REGION Network 77: Status signals
   RUNG wire#powerrail
      Contact( #TMP_xAlwaysON )
      wire#w1
      Contact( #STC_tPZD_OpCLLoop.tR.tZSW1.x0 )
      Coil( #STC_tUSER_DATA.tR.xReadyfForSwitchOn )
   END_RUNG
   RUNG wire#w1
      Contact( #STC_tPZD_OpCLLoop.tR.tZSW1.x1 )
      Contact( #STC_tPZD_OpCLLoop.tR.tZSW1.x2 )
      Coil( #STC_tUSER_DATA.tR.xReadyToMove )
   END_RUNG
   RUNG wire#w1
      Contact( #STC_tPZD_OpCLLoop.tR.tZSW1.x1 )
      Contact( #STC_tPZD_OpCLLoop.tR.tZSW1.x10 )
      Coil( #OUT_xFeedback )
   END_RUNG
   RUNG wire#w1
      Contact( #STC_tPZD_OpCLLoop.tR.tZSW1.x3 )
      wire#w2
      Coil( #OUT_xFaultPresent )
   END_RUNG
   RUNG wire#w1
      { S7_Templates := "SrcType := Int" } NE_Contact(in1 := #OUT_iRetVal, in2 := 0)
   END_RUNG wire#w2
   RUNG wire#w1
      Contact( #STC_tPZD_OpCLLoop.tR.tZSW1.x7 )
      Coil( #STC_tUSER_DATA.tR.xAlarmPresent )
   END_RUNG
   // the same network as SCL:
   #STC_tUSER_DATA.tR.xReadyfForSwitchOn := #TMP_xAlwaysON AND #STC_tPZD_OpCLLoop.tR.tZSW1.x0;
   #STC_tUSER_DATA.tR.xReadyToMove := #TMP_xAlwaysON AND #STC_tPZD_OpCLLoop.tR.tZSW1.x1 AND #STC_tPZD_OpCLLoop.tR.tZSW1.x2;
   #OUT_xFeedback := #TMP_xAlwaysON AND #STC_tPZD_OpCLLoop.tR.tZSW1.x1 AND #STC_tPZD_OpCLLoop.tR.tZSW1.x10;
   #OUT_xFaultPresent := #TMP_xAlwaysON AND (#STC_tPZD_OpCLLoop.tR.tZSW1.x3 OR (#OUT_iRetVal <> 0));
   #STC_tUSER_DATA.tR.xAlarmPresent := #TMP_xAlwaysON AND #STC_tPZD_OpCLLoop.tR.tZSW1.x7;
END_REGION

REGION Network 78: Status values
   RUNG wire#powerrail
      Contact( #TMP_xAlwaysON )
      wire#w1
      { S7_Templates := "[SrcType := DInt, DestType := Real]"; S7_GenerateENO := "TRUE" } Convert(in := #STC_tSYS_DATA.dMaxSpeed_rpm, out => #TMP_r)
      { S7_Templates := "SrcType := Real"; S7_GenerateENO := "TRUE" } Div(in1 := 16384.0, in2 := #TMP_r, out => #TMP_r)
   END_RUNG
   RUNG wire#w1
      { S7_Templates := "[SrcType := Int, DestType := DInt]"; S7_GenerateENO := "TRUE" } Convert(in := #STC_tPZD_OpCLLoop.tR.iNIST_A, out => #TMP_d)
      { S7_Templates := "[SrcType := DInt, DestType := Real]"; S7_GenerateENO := "TRUE" } Convert(in := #TMP_d, out => #TMP_rActualSpeed)
   END_RUNG
   RUNG wire#w1
      { S7_Templates := "SrcType := Real"; S7_GenerateENO := "TRUE" } Div(in1 := #TMP_rActualSpeed, in2 := #TMP_r, out => #TMP_rActualSpeed)
      { S7_Templates := "SrcType := Real"; S7_GenerateENO := "TRUE" } Mul(in1 := #TMP_rActualSpeed, in2 := #STC_tSYS_DATA.rK_rpm_mmMin, out => #TMP_rActualSpeed)
      { S7_Templates := "[SrcType := Real, DestType := DInt]"; S7_GenerateENO := "TRUE" } Trunc(in := #TMP_rActualSpeed, out => #STC_tUSER_DATA.tR.dActualSpeed_mm_min)
   END_RUNG
   // the same network as SCL:
   // ENO of a box is taken as its EN; it also drops when the box reports an error
   IF #TMP_xAlwaysON THEN
       #TMP_r := DINT_TO_REAL(#STC_tSYS_DATA.dMaxSpeed_rpm);
       #TMP_r := 16384.0 / #TMP_r;
       #TMP_d := INT_TO_DINT(#STC_tPZD_OpCLLoop.tR.iNIST_A);
       #TMP_rActualSpeed := DINT_TO_REAL(#TMP_d);
       #TMP_rActualSpeed := #TMP_rActualSpeed / #TMP_r;
       #TMP_rActualSpeed := #TMP_rActualSpeed * #STC_tSYS_DATA.rK_rpm_mmMin;
       #STC_tUSER_DATA.tR.dActualSpeed_mm_min := TRUNC(#TMP_rActualSpeed);
   END_IF;
END_REGION

REGION Network 79: #####_STATUSES_#####
END_REGION

REGION Network 80: #####_ALARMS_#####
END_REGION

REGION Network 81: Reset faults
   RUNG wire#powerrail
      Contact( #STC_tPZD_OpCLLoop.tR.tZSW1.x3 )
      Contact( #IN_xResetFaults )
      Coil( #STC_tPZD_OpCLLoop.tW.tSTW1.x7 )
   END_RUNG
   // the same network as SCL:
   #STC_tPZD_OpCLLoop.tW.tSTW1.x7 := #STC_tPZD_OpCLLoop.tR.tZSW1.x3 AND #IN_xResetFaults;
END_REGION

REGION Network 82: Fault messages
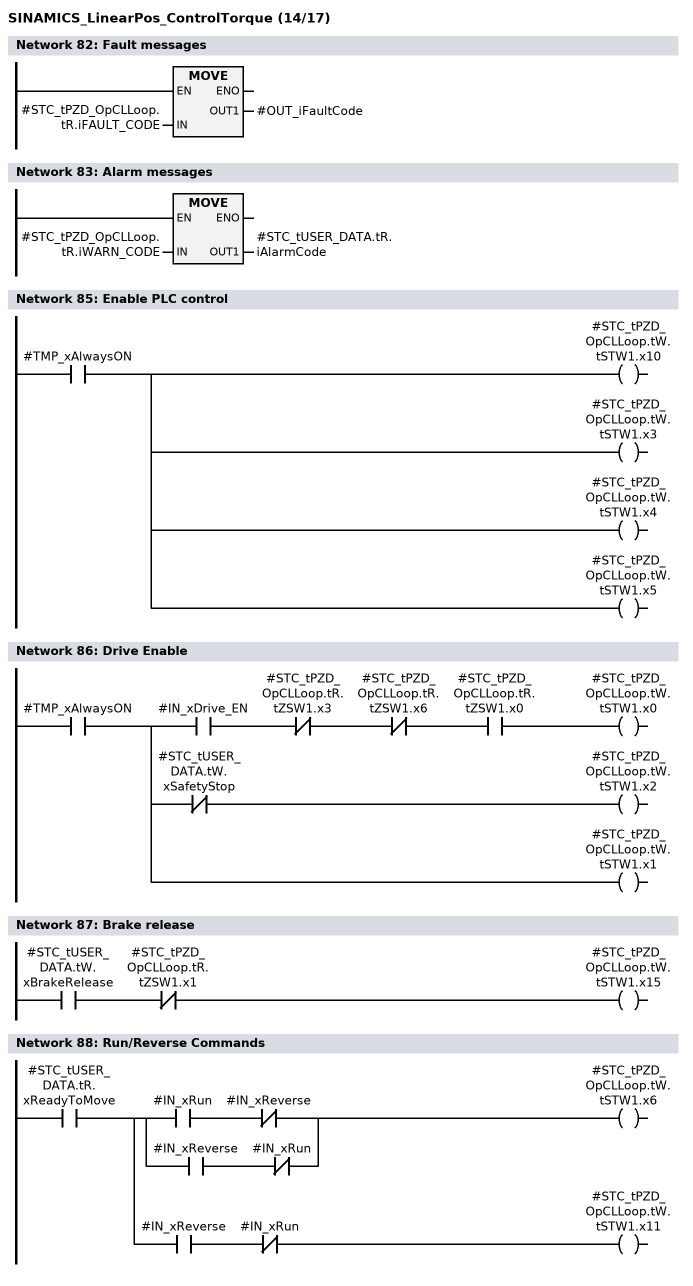
   RUNG wire#powerrail
      { S7_GenerateENO := "TRUE" } Move(in := #STC_tPZD_OpCLLoop.tR.iFAULT_CODE, out1 => #OUT_iFaultCode)
   END_RUNG
   // the same network as SCL:
   #OUT_iFaultCode := #STC_tPZD_OpCLLoop.tR.iFAULT_CODE;
END_REGION

REGION Network 83: Alarm messages
   RUNG wire#powerrail
      { S7_GenerateENO := "TRUE" } Move(in := #STC_tPZD_OpCLLoop.tR.iWARN_CODE, out1 => #STC_tUSER_DATA.tR.iAlarmCode)
   END_RUNG
   // the same network as SCL:
   #STC_tUSER_DATA.tR.iAlarmCode := #STC_tPZD_OpCLLoop.tR.iWARN_CODE;
END_REGION

REGION Network 84: #####_PHASES_&_LOGICS_#####
END_REGION

REGION Network 85: Enable PLC control
   RUNG wire#powerrail
      Contact( #TMP_xAlwaysON )
      wire#w1
      Coil( #STC_tPZD_OpCLLoop.tW.tSTW1.x10 )
   END_RUNG
   RUNG wire#w1
      Coil( #STC_tPZD_OpCLLoop.tW.tSTW1.x3 )
   END_RUNG
   RUNG wire#w1
      Coil( #STC_tPZD_OpCLLoop.tW.tSTW1.x4 )
   END_RUNG
   RUNG wire#w1
      Coil( #STC_tPZD_OpCLLoop.tW.tSTW1.x5 )
   END_RUNG
   // the same network as SCL:
   #STC_tPZD_OpCLLoop.tW.tSTW1.x10 := #TMP_xAlwaysON;
   #STC_tPZD_OpCLLoop.tW.tSTW1.x3 := #TMP_xAlwaysON;
   #STC_tPZD_OpCLLoop.tW.tSTW1.x4 := #TMP_xAlwaysON;
   #STC_tPZD_OpCLLoop.tW.tSTW1.x5 := #TMP_xAlwaysON;
END_REGION

REGION Network 86: Drive Enable
   RUNG wire#powerrail
      Contact( #TMP_xAlwaysON )
      wire#w1
      Contact( #IN_xDrive_EN )
      I_Contact( #STC_tPZD_OpCLLoop.tR.tZSW1.x3 )
      I_Contact( #STC_tPZD_OpCLLoop.tR.tZSW1.x6 )
      Contact( #STC_tPZD_OpCLLoop.tR.tZSW1.x0 )
      Coil( #STC_tPZD_OpCLLoop.tW.tSTW1.x0 )
   END_RUNG
   RUNG wire#w1
      I_Contact( #STC_tUSER_DATA.tW.xSafetyStop )
      Coil( #STC_tPZD_OpCLLoop.tW.tSTW1.x2 )
   END_RUNG
   RUNG wire#w1
      Coil( #STC_tPZD_OpCLLoop.tW.tSTW1.x1 )
   END_RUNG
   // the same network as SCL:
   #STC_tPZD_OpCLLoop.tW.tSTW1.x0 := #TMP_xAlwaysON AND #IN_xDrive_EN AND NOT #STC_tPZD_OpCLLoop.tR.tZSW1.x3 AND NOT #STC_tPZD_OpCLLoop.tR.tZSW1.x6 AND #STC_tPZD_OpCLLoop.tR.tZSW1.x0;
   #STC_tPZD_OpCLLoop.tW.tSTW1.x2 := #TMP_xAlwaysON AND NOT #STC_tUSER_DATA.tW.xSafetyStop;
   #STC_tPZD_OpCLLoop.tW.tSTW1.x1 := #TMP_xAlwaysON;
END_REGION

REGION Network 87: Brake release
   RUNG wire#powerrail
      Contact( #STC_tUSER_DATA.tW.xBrakeRelease )
      I_Contact( #STC_tPZD_OpCLLoop.tR.tZSW1.x1 )
      Coil( #STC_tPZD_OpCLLoop.tW.tSTW1.x15 )
   END_RUNG
   // the same network as SCL:
   #STC_tPZD_OpCLLoop.tW.tSTW1.x15 := #STC_tUSER_DATA.tW.xBrakeRelease AND NOT #STC_tPZD_OpCLLoop.tR.tZSW1.x1;
END_REGION

REGION Network 88: Run/Reverse Commands
   RUNG wire#powerrail
      Contact( #STC_tUSER_DATA.tR.xReadyToMove )
      wire#w1
      Contact( #IN_xRun )
      I_Contact( #IN_xReverse )
      wire#w2
      Coil( #STC_tPZD_OpCLLoop.tW.tSTW1.x6 )
   END_RUNG
   RUNG wire#w1
      Contact( #IN_xReverse )
      I_Contact( #IN_xRun )
   END_RUNG wire#w2
   RUNG wire#w1
      Contact( #IN_xReverse )
      I_Contact( #IN_xRun )
      Coil( #STC_tPZD_OpCLLoop.tW.tSTW1.x11 )
   END_RUNG
   // the same network as SCL:
   #STC_tPZD_OpCLLoop.tW.tSTW1.x6 := #STC_tUSER_DATA.tR.xReadyToMove AND ((#IN_xRun AND NOT #IN_xReverse) OR (#IN_xReverse AND NOT #IN_xRun));
   #STC_tPZD_OpCLLoop.tW.tSTW1.x11 := #STC_tUSER_DATA.tR.xReadyToMove AND #IN_xReverse AND NOT #IN_xRun;
END_REGION

REGION Network 89: #####_PARAMETERS_#####
END_REGION

REGION Network 90: Speed
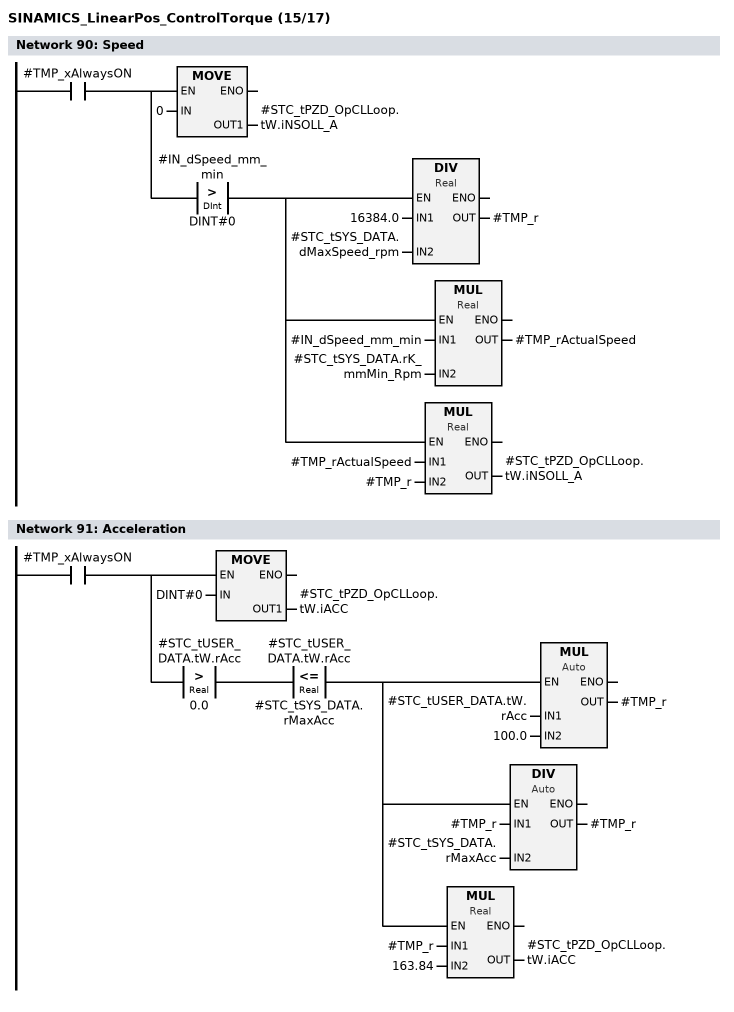
   RUNG wire#powerrail
      Contact( #TMP_xAlwaysON )
      wire#w1
      Move(in := 0, out1 => #STC_tPZD_OpCLLoop.tW.iNSOLL_A)
   END_RUNG
   RUNG wire#w1
      { S7_Templates := "SrcType := DInt" } GT_Contact(in1 := #IN_dSpeed_mm_min, in2 := DINT#0)
      wire#w2
      { S7_Templates := "SrcType := Real" } Div(in1 := 16384.0, in2 := #STC_tSYS_DATA.dMaxSpeed_rpm, out => #TMP_r)
   END_RUNG
   RUNG wire#w2
      { S7_Templates := "SrcType := Real" } Mul(in1 := #IN_dSpeed_mm_min, in2 := #STC_tSYS_DATA.rK_mmMin_Rpm, out => #TMP_rActualSpeed)
   END_RUNG
   RUNG wire#w2
      { S7_Templates := "SrcType := Real" } Mul(in1 := #TMP_rActualSpeed, in2 := #TMP_r, out => #STC_tPZD_OpCLLoop.tW.iNSOLL_A)
   END_RUNG
   // the same network as SCL:
   IF #TMP_xAlwaysON THEN #STC_tPZD_OpCLLoop.tW.iNSOLL_A := 0; END_IF;
   IF #TMP_xAlwaysON AND (#IN_dSpeed_mm_min > DINT#0) THEN
       #TMP_r := 16384.0 / #STC_tSYS_DATA.dMaxSpeed_rpm;
       #TMP_rActualSpeed := #IN_dSpeed_mm_min * #STC_tSYS_DATA.rK_mmMin_Rpm;
       #STC_tPZD_OpCLLoop.tW.iNSOLL_A := #TMP_rActualSpeed * #TMP_r;
   END_IF;
END_REGION

REGION Network 91: Acceleration
   RUNG wire#powerrail
      Contact( #TMP_xAlwaysON )
      wire#w1
      Move(in := DINT#0, out1 => #STC_tPZD_OpCLLoop.tW.iACC)
   END_RUNG
   RUNG wire#w1
      { S7_Templates := "SrcType := Real" } GT_Contact(in1 := #STC_tUSER_DATA.tW.rAcc, in2 := 0.0)
      { S7_Templates := "SrcType := Real" } LE_Contact(in1 := #STC_tUSER_DATA.tW.rAcc, in2 := #STC_tSYS_DATA.rMaxAcc)
      wire#w2
      Mul(in1 := #STC_tUSER_DATA.tW.rAcc, in2 := 100.0, out => #TMP_r)
   END_RUNG
   RUNG wire#w2
      Div(in1 := #TMP_r, in2 := #STC_tSYS_DATA.rMaxAcc, out => #TMP_r)
   END_RUNG
   RUNG wire#w2
      { S7_Templates := "SrcType := Real" } Mul(in1 := #TMP_r, in2 := 163.84, out => #STC_tPZD_OpCLLoop.tW.iACC)
   END_RUNG
   // the same network as SCL:
   IF #TMP_xAlwaysON THEN #STC_tPZD_OpCLLoop.tW.iACC := DINT#0; END_IF;
   IF #TMP_xAlwaysON AND (#STC_tUSER_DATA.tW.rAcc > 0.0) AND (#STC_tUSER_DATA.tW.rAcc <= #STC_tSYS_DATA.rMaxAcc) THEN
       #TMP_r := #STC_tUSER_DATA.tW.rAcc * 100.0;
       #TMP_r := #TMP_r / #STC_tSYS_DATA.rMaxAcc;
       #STC_tPZD_OpCLLoop.tW.iACC := #TMP_r * 163.84;
   END_IF;
END_REGION

REGION Network 92: Deceleration
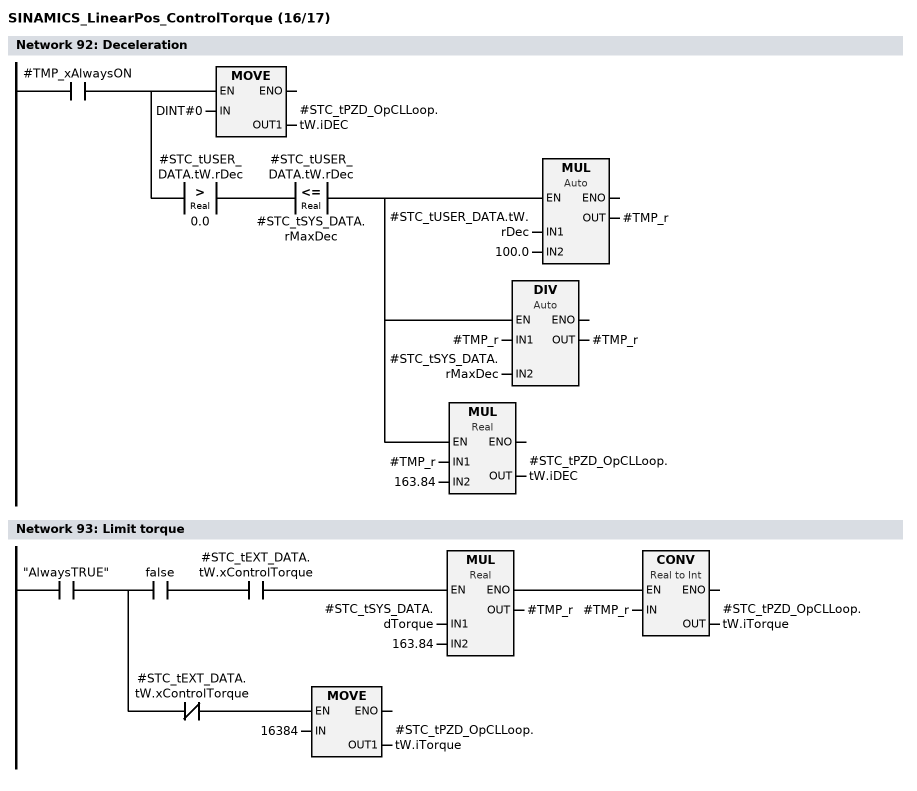
   RUNG wire#powerrail
      Contact( #TMP_xAlwaysON )
      wire#w1
      Move(in := DINT#0, out1 => #STC_tPZD_OpCLLoop.tW.iDEC)
   END_RUNG
   RUNG wire#w1
      { S7_Templates := "SrcType := Real" } GT_Contact(in1 := #STC_tUSER_DATA.tW.rDec, in2 := 0.0)
      { S7_Templates := "SrcType := Real" } LE_Contact(in1 := #STC_tUSER_DATA.tW.rDec, in2 := #STC_tSYS_DATA.rMaxDec)
      wire#w2
      Mul(in1 := #STC_tUSER_DATA.tW.rDec, in2 := 100.0, out => #TMP_r)
   END_RUNG
   RUNG wire#w2
      Div(in1 := #TMP_r, in2 := #STC_tSYS_DATA.rMaxDec, out => #TMP_r)
   END_RUNG
   RUNG wire#w2
      { S7_Templates := "SrcType := Real" } Mul(in1 := #TMP_r, in2 := 163.84, out => #STC_tPZD_OpCLLoop.tW.iDEC)
   END_RUNG
   // the same network as SCL:
   IF #TMP_xAlwaysON THEN #STC_tPZD_OpCLLoop.tW.iDEC := DINT#0; END_IF;
   IF #TMP_xAlwaysON AND (#STC_tUSER_DATA.tW.rDec > 0.0) AND (#STC_tUSER_DATA.tW.rDec <= #STC_tSYS_DATA.rMaxDec) THEN
       #TMP_r := #STC_tUSER_DATA.tW.rDec * 100.0;
       #TMP_r := #TMP_r / #STC_tSYS_DATA.rMaxDec;
       #STC_tPZD_OpCLLoop.tW.iDEC := #TMP_r * 163.84;
   END_IF;
END_REGION

REGION Network 93: Limit torque
   RUNG wire#powerrail
      Contact( "AlwaysTRUE" )
      wire#w1
      Contact( false )
      Contact( #STC_tEXT_DATA.tW.xControlTorque )
      { S7_Templates := "SrcType := Real" } Mul(in1 := #STC_tSYS_DATA.dTorque, in2 := 163.84, out => #TMP_r)
      { S7_Templates := "[SrcType := Real, DestType := Int]" } Convert(in := #TMP_r, out => #STC_tPZD_OpCLLoop.tW.iTorque)
   END_RUNG
   RUNG wire#w1
      I_Contact( #STC_tEXT_DATA.tW.xControlTorque )
      Move(in := 16384, out1 => #STC_tPZD_OpCLLoop.tW.iTorque)
   END_RUNG
   // the same network as SCL:
   IF "AlwaysTRUE" AND false AND #STC_tEXT_DATA.tW.xControlTorque THEN
       #TMP_r := #STC_tSYS_DATA.dTorque * 163.84;
       #STC_tPZD_OpCLLoop.tW.iTorque := REAL_TO_INT(#TMP_r);
   END_IF;
   IF "AlwaysTRUE" AND NOT #STC_tEXT_DATA.tW.xControlTorque THEN
       #STC_tPZD_OpCLLoop.tW.iTorque := 16384;
   END_IF;
END_REGION

REGION Network 94: ################_MOTOR_MODULE_TELEGRAMS_ENDING_#################
END_REGION

REGION Network 95 (STL): Output copy motor module
   Out:  L     #STC_tSYS_DATA.iPZD_MM;
         L     111;
         ==I;
         L     14;
         T     #TMP_iAddressLength;
         JC    WOut;
         L     #STC_tSYS_DATA.iPZD_MM;
         L     1;
         ==I;
         L     6;
         T     #TMP_iAddressLength;
         JC    WOut;

         L     19;
         JU    Err;

   WOut: NOP   0;

   //Compute destination position
         L;
         LAR1;
   //byte 1 = 10h (FIXED for S7)
         L     B#16#10;
         T     B[AR1, P#0.0];
   //byte 2 = data type
         L     B#16#4;  //4 = word
         T     B[AR1, P#1.0];
   //byte 3 & 4 = number of element
         L     #TMP_iAddressLength;  //Production data
         T     W[AR1, P#2.0];
   //byte 5 & 6 = number of DB
         L     0;  //DB production data
         T     W[AR1, P#4.0];
   //byte 7 = memory area
         L     B#16#82;  //82h = Q (Output)
         T     B[AR1, P#6.0];
   //byte 8 & 9 = address. Bit 0,1,2 of tenth byte is bit offset
   //byte 7 = address (high). Valid value = 0-7. Bit 3,4,5,6,7 always 0
         L     #STC_tSYS_DATA.iIOAddress_MM;  //Item size
         SLW   3;
         T     W[AR1, P#8.0];
         SRD   16;
         AW    16#0007;
         T     B[AR1, P#7.0];

         L     #STC_tSYS_DATA.iPZD_MM;
         L     1;
         ==I;
         JC    W1;

         CALL  BLKMOV
         ( SRCBLK  := #STC_tPZD_Pos.tW,
           RET_VAL := #TMP_iRetVal,
           DSTBLK  := #TMP_a
         );

         JU    WEnd;

   W1:   CALL  BLKMOV
         ( SRCBLK  := #STC_tPZD_OpCLLoop.tW,
           RET_VAL := #TMP_iRetVal,
           DSTBLK  := #TMP_a
         );

   WEnd: NOP   0;
END_REGION

REGION Network 96: #####_RETVAL_RESPONSE_#####
END_REGION

REGION Network 97 (STL): Initialize RetVal
         L     0;
         T     #OUT_iRetVal;
END_REGION

REGION Network 98: Warning messages
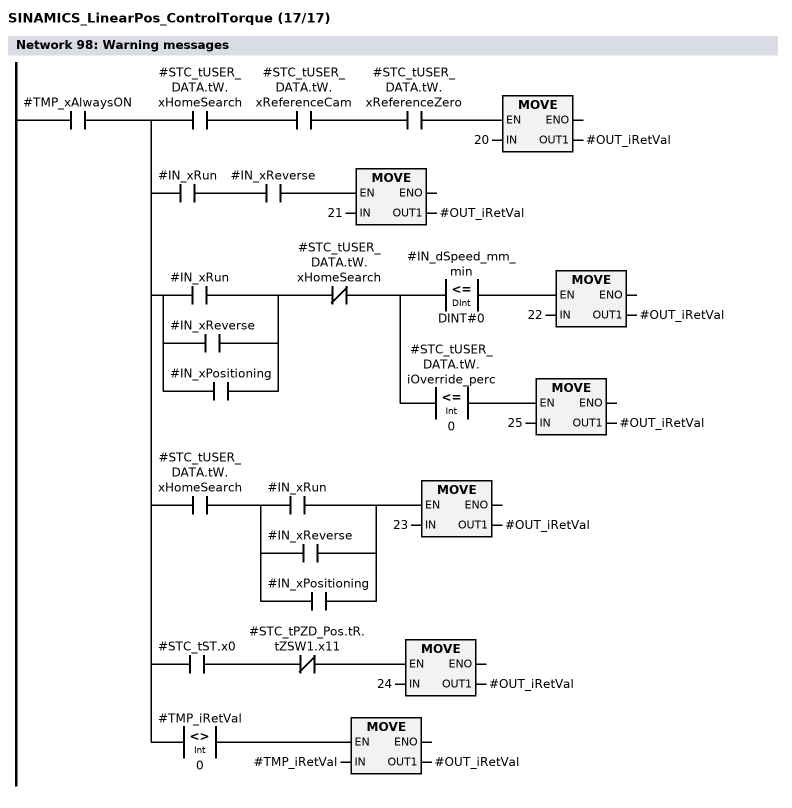
   RUNG wire#powerrail
      Contact( #TMP_xAlwaysON )
      wire#w1
      Contact( #STC_tUSER_DATA.tW.xHomeSearch )
      Contact( #STC_tUSER_DATA.tW.xReferenceCam )
      Contact( #STC_tUSER_DATA.tW.xReferenceZero )
      Move(in := 20, out1 => #OUT_iRetVal)
   END_RUNG
   RUNG wire#w1
      Contact( #IN_xRun )
      Contact( #IN_xReverse )
      Move(in := 21, out1 => #OUT_iRetVal)
   END_RUNG
   RUNG wire#w1
      Contact( #IN_xRun )
      wire#w2
      I_Contact( #STC_tUSER_DATA.tW.xHomeSearch )
      wire#w3
      { S7_Templates := "SrcType := DInt" } LE_Contact(in1 := #IN_dSpeed_mm_min, in2 := DINT#0)
      Move(in := 22, out1 => #OUT_iRetVal)
   END_RUNG
   RUNG wire#w1
      Contact( #IN_xReverse )
   END_RUNG wire#w2
   RUNG wire#w1
      Contact( #IN_xPositioning )
   END_RUNG wire#w2
   RUNG wire#w3
      { S7_Templates := "SrcType := Int" } LE_Contact(in1 := #STC_tUSER_DATA.tW.iOverride_perc, in2 := 0)
      Move(in := 25, out1 => #OUT_iRetVal)
   END_RUNG
   RUNG wire#w1
      Contact( #STC_tUSER_DATA.tW.xHomeSearch )
      wire#w4
      Contact( #IN_xRun )
      wire#w5
      Move(in := 23, out1 => #OUT_iRetVal)
   END_RUNG
   RUNG wire#w4
      Contact( #IN_xReverse )
   END_RUNG wire#w5
   RUNG wire#w4
      Contact( #IN_xPositioning )
   END_RUNG wire#w5
   RUNG wire#w1
      Contact( #STC_tST.x0 )
      I_Contact( #STC_tPZD_Pos.tR.tZSW1.x11 )
      Move(in := 24, out1 => #OUT_iRetVal)
   END_RUNG
   RUNG wire#w1
      { S7_Templates := "SrcType := Int" } NE_Contact(in1 := #TMP_iRetVal, in2 := 0)
      Move(in := #TMP_iRetVal, out1 => #OUT_iRetVal)
   END_RUNG
   // the same network as SCL:
   IF #TMP_xAlwaysON AND #STC_tUSER_DATA.tW.xHomeSearch AND #STC_tUSER_DATA.tW.xReferenceCam AND #STC_tUSER_DATA.tW.xReferenceZero THEN
       #OUT_iRetVal := 20;
   END_IF;
   IF #TMP_xAlwaysON AND #IN_xRun AND #IN_xReverse THEN #OUT_iRetVal := 21; END_IF;
   #_w1 := #TMP_xAlwaysON AND (#IN_xRun OR #IN_xReverse OR #IN_xPositioning) AND NOT #STC_tUSER_DATA.tW.xHomeSearch;
   IF #_w1 AND (#IN_dSpeed_mm_min <= DINT#0) THEN #OUT_iRetVal := 22; END_IF;
   IF #_w1 AND (#STC_tUSER_DATA.tW.iOverride_perc <= 0) THEN #OUT_iRetVal := 25; END_IF;
   IF #TMP_xAlwaysON AND #STC_tUSER_DATA.tW.xHomeSearch AND (#IN_xRun OR #IN_xReverse OR #IN_xPositioning) THEN
       #OUT_iRetVal := 23;
   END_IF;
   IF #TMP_xAlwaysON AND #STC_tST.x0 AND NOT #STC_tPZD_Pos.tR.tZSW1.x11 THEN #OUT_iRetVal := 24; END_IF;
   IF #TMP_xAlwaysON AND (#TMP_iRetVal <> 0) THEN #OUT_iRetVal := #TMP_iRetVal; END_IF;
END_REGION

REGION Network 99 (STL): Blocking messages
         JU    Rest;
   Err:  T     #OUT_iRetVal;
END_REGION

REGION Network 100 (STL): Reset input commands
   // R     #USER_DATA.W.SafetyStop
   //       R     #USER_DATA.W.FlyChange
   //       R     #USER_DATA.W.PH_Select
   //       R     #USER_DATA.W.StartCountOnHead
   //       R     #USER_DATA.W.StartCountOnTail
   //       R     #USER_DATA.W.BrakeRelease
   //       R     #USER_DATA.W.ResetCount
   //       R     #USER_DATA.W.PresetRq
   //       R     #USER_DATA.W.HomeSearch
   //       R     #USER_DATA.W.ReverseHoming
   //       R     #USER_DATA.W.ReferenceCam
   //       R     #USER_DATA.W.ReferenceZero
   //       R     #USER_DATA.W.MDI_Continue
   //       R     #USER_DATA.W.SwLimitsEnable
   //       R     #USER_DATA.W.HwLimitsEnable
   //       R     #Run
   //       R     #Reverse
   //       R     #Positioning
   // 
   //       L     L#0
   //       T     #Speed
   //       T     #USER_DATA.W.Override
   //       T     #USER_DATA.W.Target
   //       T     #USER_DATA.W.Preset
   //       T     #USER_DATA.W.Acc
   //       T     #USER_DATA.W.Dec
   Rest: NOP   0;
   //    SET
   //    R     #IN_xDrive_EN
   //    R     #IN_xResetFaults
END_REGION

REGION Network 101 (STL): Restore AR1 & AR2 value
   //    L     #TMP_dOldValue_AR1
   //    LAR1
   //    L     #TMP_dOldValue_AR2
   //    LAR2
END_REGION
END_FUNCTION_BLOCK

FUNCTION_BLOCK "SINAMICS_ClockSync"   // FB59, LAD
{ S7_Optimized_Access := 'FALSE' }
AUTHOR : Armitano
VERSION : 1.4
   VAR_INPUT
      IN_xRqSync : Bool;   // Synchronization request
   END_VAR
   VAR_OUTPUT
      OUT_xBusy : Bool;
      OUT_xDone : Bool;
      OUT_xError : Bool;
      OUT_iRetVal : Int;
   END_VAR
   VAR
      STC_tSYS_DATA : Struct   // System data
         iIOAddress_CU : Int := -1;   // Input/Output addresses for control unit
         iPosPZD_CU : Int := 1;   // Number of PZD position in SINAMICS configuration [1,2,3..]
         iDiagAddress_CU : Int;   // (NOT USED) Diagnostic addresses for control unit
      END_STRUCT;
      STC_tPROP : Struct
         xOSR_RqSync : Bool;
         xAuxBusy : Bool;
         iSyncState : Int;   // Synchronization status
         dtDateAndTimeCPU : Date_And_Time;
         dtDateOfCPU : Date;
         dtTimeOfCPU : Time_Of_Day;
      END_STRUCT;
      STC_tW_MngSysReg : Struct   // Managment system register
         tST : Struct
            xWrite_Request : Bool;
            xDone : Bool;
            xBusy : Bool;
            xError : Bool;
            xSpare4 : Bool;
            xSpare5 : Bool;
            xSpare6 : Bool;
            xSpare7 : Bool;
            ID : Hw_Io;
            dINDEX : DInt;
            uiLEN : UInt;
            dwSTATUS : DWord;
            iSpare : Int;
         END_STRUCT;
         tDATA : Struct
            wRequest_refere_RequestID : Word := W#16#102;   // (Request_referece=01 Alwais=01 )*(RequestID=02 Change Param)
            wAxis_NoOfParameters : Word := W#16#101;   // (Axis=Num.Object)(NoOfParameters=Num of parameter to change)
            wAttribute_NoOfElements : Word := W#16#1001;   // (Attribute=10 Alwais=10)(NoOfParameters=Num of subparameter to Write)
            iParameter_number : Int := 2599;   // Parameter_number=Number of the parameter
            wSubindex : Word;   // Subindex
            wFormat_NoOfValue : Word := W#16#4301;   // (Format_NoOfValue=Format 42=Word 43=Dword)(Num. of value to transfer)
            dwRegisterValue : DWord := DW#16#1;   // Register value
         END_STRUCT;
      END_STRUCT;
      STC_tWriteRecord : WRREC;
      STC_tPZD_CU : Struct   // Control unit telegram
         tR : Struct   // READ
            tZSW1 : Struct   // R2089[1].STATUS WORD 1
               x8 : Bool;   // System time synchronized
               x9 : Bool;   // Group alarm present
               x10 : Bool;   // Group fault present
               x11 : Bool;   // Safety group message present
               x12 : Bool;   // Slave sign of lifebit 0
               x13 : Bool;   // Slave sign of life bit 1
               x14 : Bool;   // Slave sign of life bit 2
               x15 : Bool;   // Slave sign of life bit 3
               x0 : Bool;   // Reserved
               x1 : Bool;   // Reserved
               x2 : Bool;   // Reserved
               x3 : Bool;   // Fault present
               x4 : Bool;   // Reserved
               x5 : Bool;   // Reserved
               x6 : Bool;   // Reserved
               x7 : Bool;   // Alarm present
            END_STRUCT;
            tE_DIGITAL : Struct   // R2089[2].DIGITAL INPUT WORD 1
               x8 : Bool;   // DI 0
               x9 : Bool;   // DI 1
               x10 : Bool;   // DI 2
               x11 : Bool;   // DI 3
               x12 : Bool;   // DI 4
               x13 : Bool;   // DI 5
               x14 : Bool;   // DI 6
               x15 : Bool;   // DI 7
               x0 : Bool;   // DI/DO 8
               x1 : Bool;   // DI/DO 9
               x2 : Bool;   // DI/DO 10
               x3 : Bool;   // DI/DO 11
               x4 : Bool;   // DI/DO 12
               x5 : Bool;   // DI/DO 13
               x6 : Bool;   // DI/DO 14
               x7 : Bool;   // DI/DO 15
            END_STRUCT;
            tE_DIGITAL_1 : Struct   // R2089[3].DIGITAL INPUT WORD 2
               x8 : Bool;   // DI 16
               x9 : Bool;   // DI 17
               x10 : Bool;   // Reserved
               x11 : Bool;   // Reserved
               x12 : Bool;   // DI 20
               x13 : Bool;   // DI 21
               x14 : Bool;   // Reserved
               x15 : Bool;   // Reserved
               x0 : Bool;   // Reserved
               x1 : Bool;   // Reserved
               x2 : Bool;   // Reserved
               x3 : Bool;   // Reserved
               x4 : Bool;   // Reserved
               x5 : Bool;   // Reserved
               x6 : Bool;   // Reserved
               x7 : Bool;   // Reserved
            END_STRUCT;
         END_STRUCT;
         tW : Struct   // WRITE
            tSTW1 : Struct   // CONTROL WORD 1
               x8 : Bool;   // Reserved
               x9 : Bool;   // Reserved
               x10 : Bool;   // P3116.Acknowledgment automatically suppressed
               x11 : Bool;   // Reserved
               x12 : Bool;   // Master sign of life bit0
               x13 : Bool;   // Master sign of life bit1
               x14 : Bool;   // Master sign of life bit2
               x15 : Bool;   // Master sign of life bit3
               x0 : Bool;   // P681.Central misuring probe, synchronizing signal source
               x1 : Bool;   // P3104.RTC real time synchronization PING
               x2 : Bool;   // Reserved
               x3 : Bool;   // Reserved
               x4 : Bool;   // Reserved
               x5 : Bool;   // Reserved
               x6 : Bool;   // Reserved
               x7 : Bool;   // P2103.Acknowledgment faults
            END_STRUCT;
            tA_DIGITAL : Struct   // DIGITAL OUTPUT WORD 1
               x8 : Bool;   // Reserved
               x9 : Bool;   // Reserved
               x10 : Bool;   // Reserved
               x11 : Bool;   // Reserved
               x12 : Bool;   // Reserved
               x13 : Bool;   // Reserved
               x14 : Bool;   // Reserved
               x15 : Bool;   // Reserved
               x0 : Bool;   // P738.CU, signal source for terminal DI/DO 8
               x1 : Bool;   // P739.CU, signal source for terminal DI/DO 9
               x2 : Bool;   // P740.CU, signal source for terminal DI/DO 10
               x3 : Bool;   // P741.CU, signal source for terminal DI/DO 11
               x4 : Bool;   // P742.CU, signal source for terminal DI/DO 12
               x5 : Bool;   // P743.CU, signal source for terminal DI/DO 13
               x6 : Bool;   // P744.CU, signal source for terminal DI/DO 14
               x7 : Bool;   // P745.CU, signal source for terminal DI/DO 15
            END_STRUCT;
            tA_DIGITAL_1 : Struct   // DIGITAL OUTPUT WORD 2
               x8 : Bool;   // Reserved
               x9 : Bool;   // Reserved
               x10 : Bool;   // Reserved
               x11 : Bool;   // Reserved
               x12 : Bool;   // Reserved
               x13 : Bool;   // Reserved
               x14 : Bool;   // Reserved
               x15 : Bool;   // Reserved
               x0 : Bool;   // Reserved
               x1 : Bool;   // Reserved
               x2 : Bool;   // Reserved
               x3 : Bool;   // Reserved
               x4 : Bool;   // Reserved
               x5 : Bool;   // Reserved
               x6 : Bool;   // Reserved
               x7 : Bool;   // Reserved
            END_STRUCT;
         END_STRUCT;
      END_STRUCT;
   END_VAR
   VAR_TEMP
      TMP_iAuxRetVal : Int;
      TMP_xAlwaysON : Bool;
      TMP_dZero : DInt;
      TMP_dIO_Pointer : DInt;
      TMP_dPZD_Pointer : DInt;
   END_VAR
BEGIN

REGION Network 1 (STL): INITIALIZATION
         SET;
         S     #TMP_xAlwaysON;
         R     #OUT_xBusy;
         R     #OUT_xDone;
         R     #OUT_xError;

         A     #STC_tPROP.xAuxBusy;
         S     #OUT_xBusy;

         L     0;
         T     #TMP_dZero;
         T     #OUT_iRetVal;

         L     #STC_tPROP.iSyncState;
         L     W#16#0;
         ==I;
         JCN   i000;
         R     #STC_tPROP.xAuxBusy;
         R     #STC_tPZD_CU.tW.tSTW1.x1;

   i000: NOP   0;
END_REGION

REGION Network 2 (STL): Copy input
   // CU Input Copy
         L     #STC_tSYS_DATA.iIOAddress_CU;
         L     0;
         <I;
         JC    NWCU;

         L     #STC_tSYS_DATA.iIOAddress_CU;
         SLW   3;
         T     #TMP_dIO_Pointer;

         L;
         T     #TMP_dPZD_Pointer;

         L     IW[ #TMP_dIO_Pointer];
         T     DIW[ #TMP_dPZD_Pointer];

         L     #TMP_dIO_Pointer;
         +     16;
         T     #TMP_dIO_Pointer;
         L     #TMP_dPZD_Pointer;
         +     16;
         T     #TMP_dPZD_Pointer;

         L     IW[ #TMP_dIO_Pointer];
         T     DIW[ #TMP_dPZD_Pointer];

         L     #TMP_dIO_Pointer;
         +     16;
         T     #TMP_dIO_Pointer;
         L     #TMP_dPZD_Pointer;
         +     16;
         T     #TMP_dPZD_Pointer;

         L     IW[ #TMP_dIO_Pointer];
         T     DIW[ #TMP_dPZD_Pointer];
END_REGION

REGION Network 3 (STL): REQUEST SYNCHRO
         A     #IN_xRqSync;
         FP    #STC_tPROP.xOSR_RqSync;
         JCN   s001;

         CALL  FILL
         ( BVAL    := #TMP_dZero,
           RET_VAL := #TMP_iAuxRetVal,
           BLK     := #STC_tW_MngSysReg
         );

         SET;
         S     #STC_tPROP.xAuxBusy;
         S     #OUT_xBusy;
         R     #STC_tPZD_CU.tW.tSTW1.x1;

         L     1;
         T     #STC_tPROP.iSyncState;
         JU    out;
   s001: NOP   0;
END_REGION

REGION Network 4 (STL): DATA FOR SETTING p3100 = 1 (UTC)
         L     #STC_tPROP.iSyncState;
         L     1;
         ==I;
         JCN   s002;

         SET;
         S     #STC_tW_MngSysReg.tST.xWrite_Request;

         L     W#16#30;  // 0x30: free choosen reference
         SLW   8;
         L     W#16#2;
         OW;
         T     #STC_tW_MngSysReg.tDATA.wRequest_refere_RequestID;
         L     #STC_tSYS_DATA.iPosPZD_CU;
         SLW   8;
         L     W#16#1;
         OW;
         T     #STC_tW_MngSysReg.tDATA.wAxis_NoOfParameters;
         L     W#16#1001;
         T     #STC_tW_MngSysReg.tDATA.wAttribute_NoOfElements;
         L     W#16#C1C;  // C1C: parameter 3100
         T     #STC_tW_MngSysReg.tDATA.iParameter_number;
         L     W#16#0;
         T     #STC_tW_MngSysReg.tDATA.wSubindex;
         L     W#16#601;
         T     #STC_tW_MngSysReg.tDATA.wFormat_NoOfValue;
         L     #STC_tSYS_DATA.iIOAddress_CU;
         T     #STC_tW_MngSysReg.tST.ID;
         L     47;
         T     #STC_tW_MngSysReg.tST.dINDEX;
         L     14;
         T     #STC_tW_MngSysReg.tST.uiLEN;

         L     W#16#1;  // 0x01: value "1"
         SLD   16;
         T     #STC_tW_MngSysReg.tDATA.dwRegisterValue;

         CALL  #STC_tWriteRecord
         ( REQ    := #STC_tW_MngSysReg.tST.xWrite_Request,
           ID     := #STC_tW_MngSysReg.tST.ID,
           INDEX  := #STC_tW_MngSysReg.tST.dINDEX,
           LEN    := #STC_tW_MngSysReg.tST.uiLEN,
           DONE   := #STC_tW_MngSysReg.tST.xDone,
           BUSY   := #STC_tW_MngSysReg.tST.xBusy,
           ERROR  := #STC_tW_MngSysReg.tST.xError,
           STATUS := #STC_tW_MngSysReg.tST.dwSTATUS,
           RECORD := #STC_tW_MngSysReg.tDATA
         );

         A     #STC_tW_MngSysReg.tST.xError;
         JCN   e002;
         S     #OUT_xError;

         L     0;
         T     #STC_tPROP.iSyncState;
         L     1;
         T     #OUT_iRetVal;
         BEU;

   e002: A     #STC_tW_MngSysReg.tST.xDone;
         JCN   s002;

         L     2;
         T     #STC_tPROP.iSyncState;

         CALL  FILL
         ( BVAL    := #TMP_dZero,
           RET_VAL := #TMP_iAuxRetVal,
           BLK     := #STC_tW_MngSysReg
         );
         JU    out;
   s002: NOP   0;
END_REGION

REGION Network 5 (STL): SET "PING" (BIT 1) IN STW1 OF CU
         L     #STC_tPROP.iSyncState;
         L     2;
         ==I;
         JCN   s003;

         SET;
         S     #STC_tPZD_CU.tW.tSTW1.x1;

         L     3;
         T     #STC_tPROP.iSyncState;
         JU    out;
   s003: NOP   0;
END_REGION

REGION Network 6 (STL): GET DATE AND TIME OF S7 CPU
         L     #STC_tPROP.iSyncState;
         L     3;
         ==I;
         JCN   s004;

         CALL  RD_LOC_T  // read clock of CPU
         ( RET_VAL := #TMP_iAuxRetVal,
           OUT     := #STC_tPROP.dtDateAndTimeCPU
         );

         CALL  T_CONV  // get date of CPU
         ( IN  := #STC_tPROP.dtDateAndTimeCPU,
           OUT := #STC_tPROP.dtDateOfCPU
         );

         CALL  T_CONV  // get time of CPU
         ( IN  := #STC_tPROP.dtDateAndTimeCPU,
           OUT := #STC_tPROP.dtTimeOfCPU
         );

         L     4;
         T     #STC_tPROP.iSyncState;
         JU    out;
   s004: NOP   0;
END_REGION

REGION Network 7 (STL): DATA FOR SETTING p3101[1]
         L     #STC_tPROP.iSyncState;
         L     4;
         ==I;
         JCN   s005;

         SET;
         S     #STC_tW_MngSysReg.tST.xWrite_Request;

         L     W#16#10;  // 0x10: free choosen reference
         SLW   8;
         L     W#16#2;
         OW;
         T     #STC_tW_MngSysReg.tDATA.wRequest_refere_RequestID;
         L     #STC_tSYS_DATA.iPosPZD_CU;
         SLW   8;
         L     W#16#1;
         OW;
         T     #STC_tW_MngSysReg.tDATA.wAxis_NoOfParameters;
         L     W#16#1001;
         T     #STC_tW_MngSysReg.tDATA.wAttribute_NoOfElements;
         L     W#16#C1D;  // C1D: parameter 3101
         T     #STC_tW_MngSysReg.tDATA.iParameter_number;
         L     W#16#1;  // 0x0001: second element of array
         T     #STC_tW_MngSysReg.tDATA.wSubindex;
         L     W#16#701;
         T     #STC_tW_MngSysReg.tDATA.wFormat_NoOfValue;
         L     #STC_tSYS_DATA.iIOAddress_CU;
         T     #STC_tW_MngSysReg.tST.ID;
         L     47;
         T     #STC_tW_MngSysReg.tST.dINDEX;
         L     16;
         T     #STC_tW_MngSysReg.tST.uiLEN;

         L     #STC_tPROP.dtDateOfCPU;  // value
         L     7305;
         +D;
         T     #STC_tW_MngSysReg.tDATA.dwRegisterValue;

         CALL  #STC_tWriteRecord
         ( REQ    := #STC_tW_MngSysReg.tST.xWrite_Request,
           ID     := #STC_tW_MngSysReg.tST.ID,
           INDEX  := #STC_tW_MngSysReg.tST.dINDEX,
           LEN    := #STC_tW_MngSysReg.tST.uiLEN,
           DONE   := #STC_tW_MngSysReg.tST.xDone,
           BUSY   := #STC_tW_MngSysReg.tST.xBusy,
           ERROR  := #STC_tW_MngSysReg.tST.xError,
           STATUS := #STC_tW_MngSysReg.tST.dwSTATUS,
           RECORD := #STC_tW_MngSysReg.tDATA
         );

         A     #STC_tW_MngSysReg.tST.xError;
         JCN   e005;
         S     #OUT_xError;

         L     0;
         T     #STC_tPROP.iSyncState;
         L     2;
         T     #OUT_iRetVal;
         BEU;

   e005: A     #STC_tW_MngSysReg.tST.xDone;
         JCN   s005;

         L     5;
         T     #STC_tPROP.iSyncState;

         CALL  FILL
         ( BVAL    := #TMP_dZero,
           RET_VAL := #TMP_iAuxRetVal,
           BLK     := #STC_tW_MngSysReg
         );
         JU    out;
   s005: NOP   0;
END_REGION

REGION Network 8 (STL): DATA FOR SETTING p3101[0]
         L     #STC_tPROP.iSyncState;
         L     5;
         ==I;
         JCN   s006;

         SET;
         S     #STC_tW_MngSysReg.tST.xWrite_Request;

         L     W#16#20;  // 0x20: free choosen reference
         SLW   8;
         L     W#16#2;
         OW;
         T     #STC_tW_MngSysReg.tDATA.wRequest_refere_RequestID;
         L     #STC_tSYS_DATA.iPosPZD_CU;
         SLW   8;
         L     W#16#1;
         OW;
         T     #STC_tW_MngSysReg.tDATA.wAxis_NoOfParameters;
         L     W#16#1001;
         T     #STC_tW_MngSysReg.tDATA.wAttribute_NoOfElements;
         L     W#16#C1D;  // C1D: parameter 3101
         T     #STC_tW_MngSysReg.tDATA.iParameter_number;
         L     W#16#0;  // 0x0000: first element of array
         T     #STC_tW_MngSysReg.tDATA.wSubindex;
         L     W#16#701;
         T     #STC_tW_MngSysReg.tDATA.wFormat_NoOfValue;
         L     #STC_tSYS_DATA.iIOAddress_CU;
         T     #STC_tW_MngSysReg.tST.ID;
         L     47;
         T     #STC_tW_MngSysReg.tST.dINDEX;
         L     16;
         T     #STC_tW_MngSysReg.tST.uiLEN;

         L     #STC_tPROP.dtTimeOfCPU;  // value
         T     #STC_tW_MngSysReg.tDATA.dwRegisterValue;

         CALL  #STC_tWriteRecord
         ( REQ    := #STC_tW_MngSysReg.tST.xWrite_Request,
           ID     := #STC_tW_MngSysReg.tST.ID,
           INDEX  := #STC_tW_MngSysReg.tST.dINDEX,
           LEN    := #STC_tW_MngSysReg.tST.uiLEN,
           DONE   := #STC_tW_MngSysReg.tST.xDone,
           BUSY   := #STC_tW_MngSysReg.tST.xBusy,
           ERROR  := #STC_tW_MngSysReg.tST.xError,
           STATUS := #STC_tW_MngSysReg.tST.dwSTATUS,
           RECORD := #STC_tW_MngSysReg.tDATA
         );

         A     #STC_tW_MngSysReg.tST.xError;
         JCN   e006;
         S     #OUT_xError;